   N128 : DINT[997] := ([0] := 1000, [1] := 1000, [2] := 1000, [3] := 1000, [4] := 1000, [5] := 1000, [6] := 1000, [30] := 6000, [42] := 6000, [54] := 6000, [66] := 6000, [78] := 6000, [90] := 6000, [96] := 200, [97] := 200, [98] := 200, [99] := 200, [100] := 100, [101] := 100, [102] := 170, [108] := 500, [109] := 1000, [110] := 1000, [111] := 800, [112] := 800, [113] := 180, [114] := 500, [126] := 1, [138] := 1000, [145] := 1, [148] := 1, [149] := 1, [157] := 1, [160] := 1, [161] := 1, [168] := 27, [169] := 27, [170] := 27, [171] := 27, [172] := 27, [173] := 27, [174] := 27, [204] := 27, [205] := 27, [206] := 27, [207] := 27, [208] := 27, [209] := 27, [210] := 27, [240] := 90, [241] := 90, [242] := 90, [243] := 90, [244] := 90, [245] := 90, [246] := 90, [252] := 12, [253] := 12, [254] := 12, [255] := 12,
        [256] := 12, [257] := 12, [258] := 12, [264] := 2, [265] := 2, [266] := 2, [267] := 2, [268] := 2, [269] := 2, [270] := 2, [276] := 1853, [277] := 1830, [278] := 1853, [279] := 1997, [280] := 1830, [281] := 2451, [282] := 2979, [288] := 6154, [289] := 6144, [290] := 6154, [291] := 6154, [292] := 6144, [293] := 6144, [294] := 6144, [300] := 6, [301] := 6, [302] := 6, [303] := 6, [304] := 6, [305] := 6, [306] := 6, [312] := 12, [313] := 12, [314] := 12, [315] := 12, [316] := 12, [317] := 12, [318] := 12, [324] := 1, [325] := 1, [326] := 1, [327] := 1, [328] := 1, [329] := 1, [330] := 1, [336] := 1, [337] := 1, [338] := 1, [339] := 1, [340] := 1, [341] := 1, [342] := 1, [348] := 1, [349] := 1, [350] := 1, [351] := 1, [352] := 1, [353] := 1, [354] := 1, [360] := 1,
        [361] := 1, [362] := 1, [363] := 1, [364] := 1, [365] := 1, [366] := 1, [372] := 1, [373] := 1, [374] := 1, [375] := 1, [376] := 1, [377] := 1, [378] := 1, [384] := 1, [385] := 1, [386] := 1, [387] := 1, [388] := 1, [389] := 1, [390] := 1, [396] := 5, [397] := 5, [398] := 5, [399] := 5, [400] := 5, [401] := 5, [402] := 5, [408] := 5, [409] := 5, [410] := 5, [411] := 5, [412] := 5, [413] := 5, [414] := 5, [437] := 100, [444] := 300, [445] := 100, [446] := 300, [447] := 300, [448] := 100, [449] := 100, [450] := 300, [457] := 1, [458] := 3, [459] := 1, [460] := 1, [462] := 3, [469] := 2, [472] := 2, [473] := 2, [486] := 1, [600] := 32, [612] := 460, [613] := 460, [614] := 460, [615] := 460, [616] := 460, [617] := 460, [618] := 460, [624] := 84,
        [625] := 84, [626] := 84, [627] := 84, [628] := 84, [629] := 84, [630] := 84, [636] := 370, [637] := 370, [638] := 370, [639] := 370, [640] := 370, [641] := 370, [642] := 370, [648] := 16384, [649] := 10922, [651] := 10922, [652] := 8745, [653] := 8745, [654] := 21845, [673] := 2048, [677] := 1639, [678] := 4096, [689] := 1091, [690] := 1259, [701] := 390, [702] := 1209, [709] := 340, [713] := 584, [714] := 735, [721] := 586, [725] := 914, [726] := 1021, [733] := 689, [737] := 1074, [738] := 1256, [745] := 280, [749] := 375, [750] := 1218, [756] := 3165, [757] := 5914, [758] := 5918, [759] := 5845, [760] := 4082, [761] := 5933, [762] := 5750, [768] := 42, [769] := 37, [770] := 43, [771] := 34, [772] := 52, [773] := 51, [774] := 58, [780] := 5, [781] := 10, [782] := 10, [783] := 40, [784] := 33, [785] := 10, [786] := 10, [792] := 5,
        [793] := 10, [794] := 10, [795] := 40, [796] := 33, [797] := 10, [798] := 10, [804] := 10, [805] := 33, [806] := 2, [807] := 43, [808] := 2, [809] := 22, [810] := 7, [816] := 5, [817] := 2, [818] := 10, [819] := 40, [820] := 7, [821] := 3, [822] := 2, [828] := 10, [829] := 33, [830] := 2, [831] := 43, [832] := 10, [833] := 10, [834] := 7, [840] := 7, [841] := 6, [842] := 2, [843] := 1, [844] := 10, [845] := 1, [846] := 1, [852] := 8, [853] := 8, [854] := 4, [855] := 2, [856] := 11, [857] := 2, [858] := 2, [864] := 13828, [865] := 10922, [876] := 3631, [877] := -28913, [878] := 3596, [880] := 3788, [891] := 1, [892] := 32, [893] := 1, [894] := 1, [912] := 83, [913] := 83, [914] := 18, [915] := 83, [917] := 83, [918] := 83, [924] := 12, [925] := 12, [926] := 6,
        [927] := 12, [928] := 6, [929] := 12, [930] := 12, [936] := 6, [937] := 6, [938] := 10, [939] := 2, [940] := 10, [941] := 6, [942] := 10, [948] := 8, [949] := 8, [950] := 11, [951] := 6, [952] := 11, [953] := 8, [954] := 11, [990] := 120, [991] := -32768, [994] := 127, [996] := 127);
        [906].1   // DEVICENET No. 1 crusher Drive Operating
        [906].7   // DEVICENET No. 1 crusher Drive faulted
        [912].6   // DEVICENET No. 1 crusher SS2 ON
        [912].7   // DEVICENET No. 1 crusher SS1 ON
   N12_HOST : INT[1000] := ([0] := 1, [1] := 650, [2] := 233, [3] := 15, [4] := 7653, [6] := 32, [7] := 31); {produced}
   N13 : DINT[48];
   N14 : DINT[1000];
        [0]   // Scanner 5 Tracking File
        [60]   // MB --> M2 CLX
        [61]   // MB --> M2 CLX
        [62]   // MB --> M2 CLX
        [63]   // MB --> M2 CLX
        [64]   // MB --> M2 CLX
        [65]   // MB --> M2 CLX
        [66]   // MB --> M2 CLX
        [67]   // MB --> M2 CLX
        [68]   // MB --> M2 CLX
        [69]   // MB --> M2 CLX
        [70]   // MB --> M2 CLX
        [71]   // MB --> M2 CLX
        [72]   // MB --> M2 CLX
        [73]   // MB --> M2 CLX
        [74]   // MB --> M2 CLX
        [75]   // MB --> M2 CLX
        [76]   // MB --> M2 CLX
        [77]   // MB --> M2 CLX
        [78]   // MB --> M2 CLX
        [79]   // MB --> M2 CLX
        [80]   // MB --> M2 CLX TD MMI Zone 2 South Skew Adjustment
        [81]   // MB --> M2 CLX TD MMI Zone 3 South Skew Adjustment
        [82]   // MB --> M2 CLX TD MMI Zone 4 South Skew Adjustment
        [83]   // MB --> M2 CLX TD MMI Zone 5 South Skew Adjustment
   N14_HOST : INT[1000]; {produced}
   N15 : DINT[1000];
   N16 : DINT[48];
   N163 : DINT[5] := ([0] := 65520, [1] := 64, [3] := 3072);
        [0]   // CROSS BREAK ZONE 3 Cross break Bit Shift 0in.--31in.
        [1]   // CROSS BREAK ZONE 3 Cross break Bit Shift 32in.--63in.
        [2]   // CROSS BREAK ZONE 3 Cross break Bit Shift 64in.in.--95in.
        [3]   // CROSS BREAK ZONE 3 Cross break Bit Shift 96in.--127in.
        [4]   // CROSS BREAK ZONE 3 Cross break Bit Shift 128in.--159in.
   N164 : DINT[3] := ([0] := 64);
        [0]   // CROSS BREAK ZONE 3 Cross break Bit Shift Compare for Sponge Roll
   N17 : DINT[1000];
        [0]   // Scanner 4 Tracking File
   N173 : DINT[360] := ([0] := 2440, [1] := 1000, [2] := 1000, [3] := 1000, [4] := 1000, [5] := 2440, [6] := 1000, [7] := 1000, [8] := 1000, [12] := 2440, [17] := 2440, [24] := 2440, [29] := 2440, [36] := 4950, [37] := 5010, [38] := 5010, [39] := 5010, [40] := 5010, [41] := 4950, [42] := 5010, [43] := 5010, [44] := 5010, [96] := 90, [97] := 90, [98] := 90, [99] := 90, [100] := 90, [101] := 90, [102] := 90, [103] := 90, [104] := 90, [108] := 90, [109] := 90, [110] := 90, [111] := 90, [112] := 90, [113] := 90, [114] := 90, [115] := 90, [116] := 90, [120] := 2440, [121] := 1000, [122] := 1000, [123] := 1000, [124] := 1000, [125] := 2440, [126] := 1000, [127] := 1000, [128] := 1000, [132] := 2440, [137] := 2440, [144] := 2440, [149] := 2440, [156] := 4950, [157] := 3345, [158] := 3345, [159] := 3345, [160] := 3345, [161] := 4950, [162] := 3345,
        [163] := 3345, [164] := 3345, [216] := 90, [217] := 90, [218] := 90, [219] := 90, [220] := 90, [221] := 90, [222] := 90, [223] := 90, [224] := 90, [228] := 90, [229] := 90, [230] := 90, [231] := 90, [232] := 90, [233] := 90, [234] := 90, [235] := 90, [236] := 90, [240] := 2440, [241] := 1000, [242] := 1000, [243] := 1000, [244] := 1000, [245] := 2440, [246] := 1000, [247] := 1000, [248] := 1000, [252] := 2440, [257] := 2440, [264] := 2440, [269] := 2440, [276] := 4950, [277] := 3900, [278] := 3900, [279] := 3900, [280] := 3900, [281] := 4950, [282] := 3900, [283] := 3900, [284] := 3900, [336] := 90, [337] := 90, [338] := 90, [339] := 90, [340] := 90, [341] := 90, [342] := 90, [343] := 90, [344] := 90, [348] := 90, [349] := 90, [350] := 90, [351] := 90, [352] := 90, [353] := 90, [354] := 90, [355] := 90, [356] := 90);
   N174 : DINT[360] := ([0] := 1000, [1] := 1000, [36] := 5010, [37] := 5010, [96] := 90, [97] := 90, [108] := 90, [109] := 90, [120] := 1000, [121] := 1000, [156] := 3345, [157] := 3345, [216] := 90, [217] := 90, [228] := 90, [229] := 90, [240] := 1000, [241] := 1000, [276] := 3900, [277] := 3900, [336] := 90, [337] := 90, [348] := 90, [349] := 90);
   N177 : DINT[5] := ([1] := 1, [2] := 80);
   N177_0 : ALIAS FOR N177[0];
   N178 : DINT[600] := ([0] := 1000, [1] := 1000, [2] := 1000, [3] := 1000, [4] := 1000, [5] := 2440, [6] := 1000, [7] := 1000, [8] := 1000, [12] := 5064, [17] := 2440, [29] := 2440, [36] := 6000, [37] := 5010, [38] := 5010, [39] := 5010, [40] := 5010, [41] := 4950, [42] := 5010, [43] := 5010, [44] := 5010, [96] := 100, [97] := 90, [98] := 90, [99] := 90, [100] := 90, [101] := 90, [102] := 90, [103] := 90, [104] := 90, [108] := 300, [109] := 90, [110] := 90, [111] := 90, [112] := 90, [113] := 90, [114] := 90, [115] := 90, [116] := 90, [168] := 27, [204] := 27, [240] := 60, [241] := 90, [242] := 90, [243] := 90, [244] := 90, [245] := 90, [246] := 90, [247] := 90, [248] := 90, [249] := 90, [250] := 90, [251] := 90, [252] := 12, [253] := 12, [254] := 12, [255] := 12, [256] := 12, [257] := 12, [258] := 12,
        [259] := 12, [260] := 12, [261] := 12, [262] := 12, [263] := 12, [264] := 2, [265] := 2, [266] := 2, [267] := 2, [268] := 2, [269] := 2, [270] := 2, [271] := 2, [272] := 2, [273] := 2, [274] := 2, [275] := 2, [276] := 4710, [277] := 1853, [278] := 1853, [279] := 1853, [280] := 1853, [281] := 1853, [282] := 1853, [283] := 1853, [284] := 1853, [285] := 1853, [286] := 1853, [287] := 1853, [288] := 6144, [289] := 6154, [290] := 6154, [291] := 6154, [292] := 6154, [293] := 6154, [294] := 6154, [295] := 6154, [296] := 6154, [297] := 6154, [298] := 6154, [299] := 6154, [300] := 6, [301] := 6, [302] := 6, [303] := 6, [304] := 6, [305] := 6, [306] := 6, [307] := 6, [308] := 6, [309] := 6, [310] := 6, [311] := 6, [312] := 12, [313] := 12, [314] := 12, [315] := 12, [316] := 12, [317] := 12, [318] := 12,
        [319] := 12, [320] := 12, [321] := 12, [322] := 12, [323] := 12, [324] := 1, [325] := 1, [326] := 1, [327] := 1, [328] := 1, [329] := 1, [330] := 1, [331] := 1, [332] := 1, [333] := 1, [334] := 1, [335] := 1, [336] := 1, [337] := 1, [338] := 1, [339] := 1, [340] := 1, [341] := 1, [342] := 1, [343] := 1, [344] := 1, [345] := 1, [346] := 1, [347] := 1, [348] := 1, [349] := 1, [350] := 1, [351] := 1, [352] := 1, [353] := 1, [354] := 1, [355] := 1, [356] := 1, [357] := 1, [358] := 1, [359] := 1, [360] := 1, [361] := 1, [362] := 1, [363] := 1, [364] := 1, [365] := 1, [366] := 1, [367] := 1, [368] := 1, [369] := 1, [370] := 1, [371] := 1, [372] := 1, [373] := 1, [374] := 1, [375] := 1, [376] := 1, [377] := 1, [378] := 1,
        [379] := 1, [380] := 1, [381] := 1, [382] := 1, [383] := 1, [384] := 1, [385] := 1, [386] := 1, [387] := 1, [388] := 1, [389] := 1, [390] := 1, [391] := 1, [392] := 1, [393] := 1, [394] := 1, [395] := 1, [396] := 5, [397] := 5, [398] := 5, [399] := 5, [400] := 5, [401] := 5, [402] := 5, [403] := 5, [404] := 5, [405] := 5, [406] := 5, [407] := 5, [408] := 5, [409] := 5, [410] := 5, [411] := 5, [412] := 5, [413] := 5, [414] := 5, [415] := 5, [416] := 5, [417] := 5, [418] := 5, [419] := 5, [432] := 300, [433] := 300, [434] := 300, [435] := 300, [436] := 300, [437] := 300, [438] := 300, [439] := 300, [440] := 300, [441] := 300, [442] := 300, [443] := 300, [444] := 300, [445] := 300, [446] := 300, [447] := 300, [448] := 300, [449] := 300, [450] := 300,
        [451] := 300, [452] := 300, [453] := 300, [454] := 300, [455] := 300, [457] := 2, [458] := 2, [459] := 2, [460] := 2, [461] := 2, [462] := 2, [463] := 2, [464] := 2, [465] := 2, [466] := 2, [467] := 2);
        [12]   // APC Frequency Setpoint for Drive Freq 1 [Hz * 100]
   N179 : DINT[600] := ([0] := 1000, [1] := 1000, [2] := 1000, [3] := 1000, [4] := 1000, [5] := 1000, [6] := 1000, [12] := 3000, [13] := 3000, [14] := 3000, [15] := 3000, [16] := 1816, [17] := 1816, [18] := 6000, [30] := 6000, [42] := 6000, [54] := 6000, [66] := 6000, [78] := 6000, [90] := 6000, [96] := 200, [97] := 200, [98] := 200, [99] := 200, [100] := 200, [101] := 100, [102] := 170, [108] := 500, [109] := 500, [110] := 500, [111] := 500, [112] := 500, [113] := 500, [114] := 500, [126] := 1, [138] := 1000, [168] := 27, [169] := 27, [170] := 27, [171] := 27, [172] := 27, [173] := 27, [174] := 27, [204] := 27, [205] := 27, [206] := 27, [207] := 27, [208] := 27, [209] := 27, [210] := 27, [240] := 90, [241] := 90, [242] := 90, [243] := 90, [244] := 90, [245] := 90, [246] := 90, [247] := 90, [248] := 90, [249] := 90,
        [250] := 90, [251] := 90, [252] := 12, [253] := 12, [254] := 12, [255] := 12, [256] := 12, [257] := 12, [258] := 12, [259] := 12, [260] := 12, [261] := 12, [262] := 12, [263] := 12, [264] := 2, [265] := 2, [266] := 2, [267] := 2, [268] := 2, [269] := 2, [270] := 2, [271] := 2, [272] := 2, [273] := 2, [274] := 2, [275] := 2, [276] := 1853, [277] := 1853, [278] := 1853, [279] := 1853, [280] := 1853, [281] := 1853, [282] := 2979, [283] := 1853, [284] := 1853, [285] := 1853, [286] := 1853, [287] := 1853, [288] := 6154, [289] := 6154, [290] := 6154, [291] := 6154, [292] := 6154, [293] := 6154, [294] := 6144, [295] := 6154, [296] := 6154, [297] := 6154, [298] := 6154, [299] := 6154, [300] := 6, [301] := 6, [302] := 6, [303] := 6, [304] := 6, [305] := 6, [306] := 6, [307] := 6, [308] := 6, [309] := 6,
        [310] := 6, [311] := 6, [312] := 12, [313] := 12, [314] := 12, [315] := 12, [316] := 12, [317] := 12, [318] := 12, [319] := 12, [320] := 12, [321] := 12, [322] := 12, [323] := 12, [324] := 1, [325] := 1, [326] := 1, [327] := 1, [328] := 1, [329] := 1, [330] := 1, [331] := 1, [332] := 1, [333] := 1, [334] := 1, [335] := 1, [336] := 1, [337] := 1, [338] := 1, [339] := 1, [340] := 1, [341] := 1, [342] := 1, [343] := 1, [344] := 1, [345] := 1, [346] := 1, [347] := 1, [348] := 1, [349] := 1, [350] := 1, [351] := 1, [352] := 1, [353] := 1, [354] := 1, [355] := 1, [356] := 1, [357] := 1, [358] := 1, [359] := 1, [360] := 1, [361] := 1, [362] := 1, [363] := 1, [364] := 1, [365] := 1, [366] := 1, [367] := 1, [368] := 1, [369] := 1,
        [370] := 1, [371] := 1, [372] := 1, [373] := 1, [374] := 1, [375] := 1, [376] := 1, [377] := 1, [378] := 1, [379] := 1, [380] := 1, [381] := 1, [382] := 1, [383] := 1, [384] := 1, [385] := 1, [386] := 1, [387] := 1, [388] := 1, [389] := 1, [390] := 1, [391] := 1, [392] := 1, [393] := 1, [394] := 1, [395] := 1, [396] := 5, [397] := 5, [398] := 5, [399] := 5, [400] := 5, [401] := 5, [402] := 5, [403] := 5, [404] := 5, [405] := 5, [406] := 5, [407] := 5, [408] := 5, [409] := 5, [410] := 5, [411] := 5, [412] := 5, [413] := 5, [414] := 5, [415] := 5, [416] := 5, [417] := 5, [418] := 5, [419] := 5, [432] := 300, [433] := 300, [434] := 300, [435] := 300, [436] := 300, [437] := 300, [438] := 300, [439] := 300, [440] := 300, [441] := 300,
        [442] := 300, [443] := 300, [444] := 300, [445] := 300, [446] := 300, [447] := 300, [448] := 300, [449] := 300, [450] := 300, [451] := 300, [452] := 300, [453] := 300, [454] := 300, [455] := 300, [462] := 2);
        [12]   // Brush 1 and 2 speed DEVICENET Conveyor 1 Speed setpnt 1 ** channel b **
        [13]   // DEVICENET Conveyor 2 Speed setpnt 1 ** channel b **
        [14]   // DEVICENET Conveyor 3 Speed setpnt 1 ** channel b **
        [15]   // DEVICENET Conveyor 4 Speed setpnt 1 ** channel b **
        [16]   // DEVICENET Conveyor 5 Speed setpnt 1 ** channel b **
        [17]   // DEVICENET Conveyor 6 Speed setpnt 1 ** channel b **
        [18]   // DEVICENET Conveyor 7 Speed setpnt 1 ** channel b **
        [30]   // DEVICENET Conveyor 7 Speed setpnt 2 ** channel b **
   N18 : DINT[1000];
   N184 : DINT[50] := ([0] := 2, [1] := 1, [2] := 2, [3] := 3, [4] := 4, [5] := 5, [6] := 6, [7] := 100, [8] := 101, [9] := 2, [11] := 900, [12] := 660, [14] := 456, [16] := 12, [17] := 47, [18] := 107, [19] := 1, [20] := 8, [21] := 171, [22] := 172, [23] := 173, [24] := 174, [25] := 175, [26] := 176, [27] := 145, [28] := 146, [29] := 128, [30] := 6, [31] := 906, [32] := 666, [34] := 462, [36] := 18, [37] := 570, [39] := 127, [49] := 64);
   N184_1 : ALIAS FOR N184[1];
   N184_10 : ALIAS FOR N184[10];
   N184_11 : ALIAS FOR N184[11];
   N184_12 : ALIAS FOR N184[12];
   N184_14 : ALIAS FOR N184[14];
   N184_16 : ALIAS FOR N184[16];
   N184_2 : ALIAS FOR N184[2];
   N184_21 : ALIAS FOR N184[21];
   N184_22 : ALIAS FOR N184[22];
   N184_23 : ALIAS FOR N184[23];
   N184_24 : ALIAS FOR N184[24];
   N184_25 : ALIAS FOR N184[25];
   N184_26 : ALIAS FOR N184[26];
   N184_3 : ALIAS FOR N184[3];
   N184_30 : ALIAS FOR N184[30];
   N184_31 : ALIAS FOR N184[31];
   N184_32 : ALIAS FOR N184[32];
   N184_34 : ALIAS FOR N184[34];
   N184_36 : ALIAS FOR N184[36];
   N184_4 : ALIAS FOR N184[4];
   N184_5 : ALIAS FOR N184[5];
   N184_6 : ALIAS FOR N184[6];
   N188 : DINT[500] := ([4] := 256, [6] := 3848, [8] := 1792, [10] := 256, [12] := 256, [14] := 1280, [16] := 256, [20] := 256, [28] := 256);
        [0]   // I/O STATUS FILE: Rack 0 FAULT/PRESENT BITS
        [1]   // I/O STATUS FILE: Rack 0 INHIBIT/RESET BITS
        [2]   // I/O STATUS FILE: Rack 1 FAULT/PRESENT BITS
        [3]   // I/O STATUS FILE: Rack 1 INHIBIT/RESET BITS
        [4]   // I/O STATUS FILE: Rack 2 FAULT/PRESENT BITS
        [6]   // I/O STATUS FILE: Rack 3 FAULT/PRESENT BITS
        [20].0   // I/O STATUS FILE: Rack 12 Group 0 FAULT
        [20].1   // I/O STATUS FILE: Rack 12 Group 2 FAULT
        [20].2   // I/O STATUS FILE: Rack 12 Group 4 FAULT
        [20].3   // I/O STATUS FILE: Rack 12 Group 6 FAULT
   N189 : DINT[40] := ([0] := -24819, [1] := 22586, [2] := -29699, [6] := -5625, [7] := -8126, [9] := 12276, [11] := 1, [12] := 11397, [13] := 21096, [14] := 5477, [15] := 11642, [16] := 11465, [18] := 45, [19] := 19110);
   N19 : DINT[48];
   N195 : DINT[50] := ([0] := 158, [1] := -4320, [2] := 7472, [3] := 6225, [4] := 7472, [5] := 6195, [7] := 30, [8] := 158, [9] := -6342, [13] := 2042, [14] := 6963, [15] := 8710, [16] := 31474, [17] := -27661, [18] := -3913, [19] := -11983, [20] := -2995, [21] := 19794, [26] := -1, [27] := -935, [33] := 2, [36] := -26, [37] := -27966, [38] := -29, [39] := 23316, [40] := -19, [41] := 17034, [44] := 4560, [46] := -17380, [47] := -19631, [48] := -30124, [49] := 3183);
   N20 : DINT[1000];
        [0]   // Scanner 4 Tracking File
   N21 : DINT[1000];
   N22 : DINT[48];
   N23 : DINT[1000];
        [0]   // Scanner 3 Tracking File
   N24 : DINT[1000];
   N25 : DINT[48];
   N250 : DINT[50] := ([30] := 1, [31] := 300, [32] := 768, [33] := 768, [34] := 300);
        [30].0   // temp test
   N251 : DINT[999];
        [900]   // DATA BITS READ BY THE WASHER PLC
        [900].0   // CITRIC ACID WASHER SOLENOID VALVE ON BIT TO WASHER PLC
        [901]   // DATA BITS WRITTEN FROM THE WASHER PLC
        [901].0   // CITRIC ACID WASHER OK BIT FROM WASHER PLC
   N26 : DINT[1000] := ([41] := 14);
        [0]   // Scanner 3 Tracking File
   N27 : DINT[1000];
   N28 : DINT[997] := ([990] := 7, [992] := 7, [993] := 7, [994] := 7, [996] := 23);
   N29 : DINT[1000];
        [0]   // Scanner 2 Tracking File
   N30 : DINT[1000];
   N31 : DINT[49];
   N32 : DINT[1000];
        [0]   // Scanner 2 Tracking File
   N33 : DINT[1000];
   N34 : DINT[48];
   N35 : DINT[1000];
        [0]   // Scanner 1 Tracking File
   N36 : DINT[1000];
   N37 : DINT[48];
   N38 : DINT[1000];
        [0]   // Scanner 1 Tracking File
   N39 : DINT[1000];
   N40 : DINT[48];
   N42 : DINT[89] := ([2] := 3, [3] := 16, [4] := 4101, [5] := 409, [6] := 600, [8] := 10, [12] := 20, [25] := 8, [29] := 1, [30] := 2, [34] := 1, [71] := 80, [73] := 302, [74] := 854, [76] := 5, [77] := 1, [78] := 136, [80] := 10, [81] := 297, [82] := 826, [85] := 1, [86] := 136);
        [1].5   // PC01 New Data Acknowledge
        [1].6   // PC03 New Data Acknowledge
        [1].7   // PC02 New Data Acknowledge
        [1].8   // PC00 Load Preset-
        [1].9   // PC01 Load Preset-
        [1].10   // PC02 Load Preset-
        [1].11   // PC03 Load Preset-
        [1].12   // Not Used
        [1].13   // Not Used
        [1].14   // Not Used
        [1].15   // VHSC Data Representation Mode 0 = Binary 1 = BCD
        [2]   // Word 2 VHSC BTW Data
        [2].0   // Output 00 Enable
        [2].1   // Output 01 Enable
        [2].2   // Output 02 Enable
        [2].3   // Output 03 Enable
        [2].4   // Output 04 Enable
        [2].5   // Output 05 Enable
        [2].6   // Output 06 Enable
        [2].7   // Output 07 Enable
        [2].8   // Output 00 Force
        [2].9   // Output 01 Force
        [2].10   // Output 02 Force
        [2].11   // Output 03 Force
        [2].12   // Output 04 Force
        [2].13   // Output 05 Force
        [2].14   // Output 06 Force
        [2].15   // Output 07 Force
        [3]   // Mode Bits For Counters 0 and 1 ** Default ** ** Used **
        [4].12   // VHSC Counter 3 Gate Mode Bit #1
        [4].14   // VHSC Counter 3 Gate Mode Bit #3
        [5]   // PC00 Rollover Value MSD
        [6]   // PC00 Rollover Value LSD
        [7]   // PC01 Rollover Value MSD
        [8]   // PC01 Rollover Value LSD
        [9]   // PC02 Rollover Value MSD
        [10]   // PC02 Rollover Value LSD
        [11]   // PC03 Rollover Value LSD
        [12]   // PC03 Rollover Value LSD
        [13]   // PC00 Preset Value MSD
        [14]   // PC00 Preset Value LSD
        [15]   // PC01 Preset Value MSD
        [16]   // PC01 Preset Value LSD
        [17]   // PC02 Preset Value MSD
        [18]   // PC02 Preset Value LSD
        [19]   // PC03 Preset Value LSD
        [21]   // Counter 0 Sample Period X 10mS
        [22]   // Counter 1 Sample Period X 10mS
        [23]   // Counter 2 Sample Period X 10mS
        [24]   // Counter 3 Sample Period X 10mS
        [25]   // *************** * Output 00 ** * Mapping ** * Bits ** ***************
        [25].0   // Output 00 Output/Counter Mapping Bits PC00
        [25].1   // Output 00 Output/Counter Mapping Bits PC01
        [25].2   // Output 00 Output/Counter Mapping Bits PC02
        [25].3   // Output 00 Output/Counter Mapping Bits PC03
        [26]   // Output 00 ON VALUE MSD
        [27]   // Output 00 ON VALUE LSD
        [28]   // Output 00 OFF VALUE MSD
        [29]   // Output 00 OFF VALUE LSD
        [30]   // *************** * Output 01 ** * Mapping ** * Bits ** ***************
        [30].0   // Output 01 Output/Counter Mapping Bits PC00
        [30].1   // Output 01 Output/Counter Mapping Bits PC01
        [30].2   // Output 01 Output/Counter Mapping Bits PC02
        [30].3   // Output 01 Output/Counter Mapping Bits PC03
        [31]   // Output 01 ON VALUE MSD
        [32]   // Output 01 ON VALUE LSD
        [33]   // Output 01 OFF VALUE MSD
        [34]   // Output 01 OFF VALUE LSD
        [35]   // *************** * Output 02 ** * Mapping ** * Bits ** ***************
        [36]   // Output 02 ON VALUE MSD
        [37]   // Output 02 ON VALUE LSD
        [38]   // Output 02 OFF VALUE MSD
        [39]   // Output 02 OFF VALUE LSD
        [40]   // *************** * Output 03 ** * Mapping ** * Bits ** ***************
        [45]   // *************** * Output 04 ** * Mapping ** * Bits ** ***************
        [46]   // Output 04 ON VALUE MSD
        [47]   // Output 04 ON VALUE LSD
        [48]   // Output 04 OFF VALUE MSD
        [49]   // Output 04 OFF VALUE LSD
        [50]   // *************** * Output 05 ** * Mapping ** * Bits ** ***************
        [55]   // *************** * Output 06 ** * Mapping ** * Bits ** ***************
        [56]   // Output 06 ON VALUE MSD
        [57]   // Output 06 ON VALUE LSD
        [58]   // Output 06 OFF VALUE MSD
        [59]   // Output 06 OFF VALUE LSD
        [60]   // *************** * Output 07 ** * Mapping ** * Bits ** ***************
        [61]   // Output 07 ON VALUE MSD
        [62]   // Output 07 ON VALUE LSD
        [63]   // Output 07 OFF VALUE MSD
        [64]   // Output 07 OFF VALUE LSD
        [71].0   // VHSC Configured Bit
        [72].0   // 1 M Sync Pulse (VHSC Output 0)
        [87]   // VHSC Counter 3 Stored Count MSD
   N43 : DINT[240] := ([0] := -1, [2] := -1, [4] := -1, [6] := -1, [8] := -1, [10] := -1, [12] := -1, [14] := -1, [16] := -1, [18] := -1, [20] := -1, [22] := -1, [24] := -1, [26] := -1, [28] := -1, [30] := -1, [32] := -1, [34] := -1, [36] := -1, [38] := -1, [40] := -1, [42] := -1, [44] := -1, [46] := -1, [48] := -1, [50] := -1, [52] := -1, [54] := -1, [56] := -1, [58] := -1, [60] := -1, [62] := -1, [64] := -1, [66] := -1, [68] := -1, [70] := -1, [72] := -1, [74] := -1, [76] := -1, [78] := -1, [80] := -1, [82] := -1, [84] := -1, [86] := -1, [88] := -1, [90] := -1, [92] := -1, [94] := -1, [96] := -1, [98] := -1, [200] := 130, [201] := 130, [202] := 131, [203] := 297, [204] := 826, [205] := 32, [206] := 641, [207] := 34, [208] := 375338, [209] := 256,
        [210] := 2706, [211] := 16, [212] := 234, [234] := 873, [235] := 34, [236] := 375338, [237] := 32, [238] := 641);
        [209]   // Signals to Host
        [0]   // Start of Flaw Buffer
        [200]   // Flaw Head Pointer from Host
        [200].0   // Head Ptr is an odd number?
